(*//状态输出*)(*状态显示，容易造成指针容量不足*)
mov( ConveyorMotor.xEmpty AND NOT ConveyorMotor.xBusy , 0 , m_wStateWord);
mov( ConveyorMotor.xEmpty=0 , 							1 , m_wStateWord);
mov( ConveyorMotor.xBusy , 								2 , m_wStateWord);
mov( ConveyorMotor.xLimitAlarrm , 						3, 	m_wStateWord);
mov(ConveyorMotor.xOverWidthAlarm , 					4 , m_wStateWord);
mov( ConveyorMotor.xNotArriveAlarm , 					5 , m_wStateWord);
mov( ConveyorMotor.xUnloadAlarm, 						6 , m_wStateWord);
(*选择本线体后，将状态赋值给全局变量进行显示*)
mov( ConveyorMotor.diDeviceID=g_diDeviceIDSelect , m_wStateWord, g_iConveyorStatus );
END_FUNCTION_BLOCK

PROGRAM TCP
VAR
  m_ton1ReceiveHeartbeat : TON;
  m_t1RecHeartbeatCurrentTime : TIME;
  m_tonAutoClose : TON;
  m_xAutoClose : BOOL;
  m_tAutoCloseCurrentTime : TIME;
  m_tonReconnect : TON;
  m_xReconnect : BOOL;
  m_tReconnectCurrentTime : TIME;
  m_ton5ReceiveHeartbeat : TON;
  m_t5RecHeartbeatCurrentTime : TIME;
END_VAR
D220:=2;
m_tonReconnect(IN:= NOT SD1282.0 AND NOT SD1284.0 AND NOT m_xReconnect ,PT:=T#5s  ,Q:=m_xReconnect ,ET:=m_tReconnectCurrentTime);
SP_SOCOPEN(m_xReconnect  AND SD1288.A , "U0", K1 , D110 , M100);
SP_SOCSND( SM412 AND SD1282.0 , "U0" , K1 , D100, D220, M102 );
SP_SOCRCV( SD1282.0 AND SD1286.0 AND NOT M104 , "U0" , K1, D300 , D420 ,M104 );
m_tonAutoClose(IN:= SD1284.0 AND NOT SD1282.0 ,PT:=T#5s,Q:=m_xAutoClose ,ET:= m_tAutoCloseCurrentTime );
SP_SOCCLOSE( LDF(TRUE,SD1282.0) OR m_xAutoClose  , "U0" , K1, D120, M106 );
D221.F:=SM413;
m_ton1ReceiveHeartbeat(IN:=NOT LDP(TRUE, D421.F) ,PT:= t#5S ,Q:= g_xTcpFailed ,ET:= m_t1RecHeartbeatCurrentTime);
IF g_xTcpFailed THEN
	M104:=SM413;(*通讯失败有可能是接收模块没动作，重启接收模块*)
	D420:=0;
	D421:=0;
END_IF;

(*测试一下通信恢复功能*)
IF  g_xTcpFailed THEN
	SD1284.0:=SM414;
	SD414:=20;
END_IF;
END_PROGRAM

FUNCTION_BLOCK UConveyor
VAR
  iStep : INT;
END_VAR
VAR_IN_OUT
  ConveyorIOLeft : ConveyorIO;  (* U的左半边 *)
  ConveyorIORight : ConveyorIO;  (* U的右半边 *)
  ConveyorIODown : ConveyorIO;  (* U的下边一横 *)
  UConveyorIO : UConveyorIO;  (* 顶升,阻挡 *)
END_VAR
VAR
  m_xInitial : BOOL;
  m_tonCylinderOvertime : TON;  (* 气缸超时报警定时器 *)
  m_tCylinderOvertimeCurrent : TIME;
  m_tonExitBarDelay : TON;  (* 退出阻挡器延时 *)
  m_tExitBarDelay : TIME;
  m_xExitBarDelay : BOOL;
END_VAR
(*                                                                                                          
           

//*)
IF NOT m_xInitial THEN
	UConveyorIO.tSetOvertime:=T#5s;
	UConveyorIO.xExitEnable1:=1;
	UConveyorIO.xExitEnable2:=1;
	UConveyorIO.xExitEnable3:=1;
	m_xInitial:=1;
END_IF;
(*外部不用写ConveyorDown的开关，会自己根据来料的产品信息判断停哪个光电*)
IF UConveyorIO.iTask=1 AND ConveyorIODown.diDesConveyorIn=ConveyorIOLeft.diDeviceID THEN
	ConveyorIODown.xCWPresent:=ConveyorIOLeft.xCWPresent;
ELSIF UConveyorIO.iTask=1 AND ConveyorIODown.diDesConveyorIn=ConveyorIORight.diDeviceID THEN
	ConveyorIODown.xCWPresent:=ConveyorIORight.xCWPresent;
ELSE
	ConveyorIODown.xCWPresent:=ConveyorIOLeft.xCWPresent OR ConveyorIORight.xCWPresent;
END_IF;
(*这里判断什么时候直接放行，左右都不需要，也不是0，就放走*)
IF  NOT(ConveyorIODown.diDesConveyor=ConveyorIOLeft.diDeviceID 
		OR  ConveyorIODown.diDesConveyor=ConveyorIORight.diDeviceID 
		OR ConveyorIODown.diDesConveyor=0) THEN
	UConveyorIO.xPassEnable:=1;
ELSE
	UConveyorIO.xPassEnable:=0;
END_IF;	
IF g_xAuto THEN	
CASE UConveyorIO.iTask OF(*这个Task做抢占，可做LastTask保护*)
0:(*各种初始化，能自动去3*)
	ConveyorIODown.xLoad:=0;
	ConveyorIOleft.xLoad:=0;
	ConveyorIORight.xLoad:=0;
	ConveyorIODown.xUnload:=0;
	ConveyorIOLeft.xUnload:=0;
	ConveyorIORight.xUnload:=0;
	ConveyorIODown.xPutInto:=0;
	ConveyorIOLeft.xPutInto:=0;
	ConveyorIORight.xPutInto:=0;
	UConveyorIO.xExitBarCylinderRetract1:=0;
	UConveyorIO.xExitBarCylinderRetract2:=0;	
1:(*上料*)
	CASE iStep OF
	0:(*各种初始化，能自动去3*)
		ConveyorIODown.xLoad:=0;
		ConveyorIOleft.xLoad:=0;
		ConveyorIORight.xLoad:=0;
		ConveyorIODown.xUnload:=0;
		ConveyorIOLeft.xUnload:=0;
		ConveyorIORight.xUnload:=0;
		ConveyorIODown.xPutInto:=0;
		ConveyorIOLeft.xPutInto:=0;
		ConveyorIORight.xPutInto:=0;
		UConveyorIO.xExitBarCylinderRetract1:=0;
		UConveyorIO.xExitBarCylinderRetract2:=0;
		UConveyorIO.xBatteryError:=0;
		IF  NOT ConveyorIODown.xEmpty THEN
			iStep:=3;
		ELSE
			iStep:=1;
		END_IF;	
	1:(*顶升，等load*)
		IF UConveyorIO.xLiftCylinderExtendInit1 THEN
			UConveyorIO.xLiftCylinderExtend1:=1;
			UConveyorIO.xLiftCylinderRetract1:=0;
		ELSE
			UConveyorIO.xLiftCylinderExtend1:=0;
			UConveyorIO.xLiftCylinderRetract1:=1;
		END_IF;
		IF UConveyorIO.xLiftCylinderExtendInit2 THEN
			UConveyorIO.xLiftCylinderExtend2:=1;
			UConveyorIO.xLiftCylinderRetract2:=0;
			ELSE
			UConveyorIO.xLiftCylinderExtend2:=0;
			UConveyorIO.xLiftCylinderRetract2:=1;
		END_IF;
		IF 	((UConveyorIO.xLiftCylinderExtendInit1 AND UConveyorIO.xLiftCylinderExtendDetect1)
				OR (NOT UConveyorIO.xLiftCylinderExtendInit1 AND UConveyorIO.xLiftCylinderRetractDetect1))
			AND	((UConveyorIO.xLiftCylinderExtendInit2 AND UConveyorIO.xLiftCylinderExtendDetect2)
		   		OR (NOT UConveyorIO.xLiftCylinderExtendInit2 AND UConveyorIO.xLiftCylinderRetractDetect2))		
			AND	UConveyorIO.xEntryEnable1 THEN(*有上料请求1*)
		   	ConveyorIODown.xLoad:=1;
			iStep:=2;
		END_IF;
	2:(*Load完成*)(*去右臂时才需要阻挡放行,其他挡住*)
		UConveyorIO.xExitBarCylinderRetract1:=ConveyorIODown.diDesConveyorIn=ConveyorIORight.diDeviceID;
		IF NOT ConveyorIODown.xEmpty THEN
			ConveyorIODown.xLoad:=0;
			ConveyorIOLeft.xPutInto:=1;
			ConveyorIOright.xPutInto:=1;
			istep:=3;
		END_IF;
	3:(*顶升等Unload，这里等有了ExitEnable再顶升，因为可能有地方需要允许了再升降，比如倍速链*)
	IF (ConveyorIODown.diDesConveyor=ConveyorIOLeft.diDeviceID OR ConveyorIODown.diDesConveyor=ConveyorIORight.diDeviceID)
			AND	(UConveyorIO.xBatteryDetect1 OR UConveyorIO.xBatteryDetect2)(*在下面时检测*)
			AND UConveyorIO.xLiftCylinderRetractDetect1 AND UConveyorIO.xLiftCylinderRetractDetect2 THEN
			UConveyorIO.xBatteryError:=1;
		END_IF;	
		IF (ConveyorIODown.diDesConveyor=ConveyorIOLeft.diDeviceID AND UConveyorIO.xExitEnable2 AND NOT UConveyorIO.xBatteryError)THEN
			IF UConveyorIO.xLiftCylinderExtendInit1 THEN
				UConveyorIO.xLiftCylinderExtend1:=0;
				UConveyorIO.xLiftCylinderRetract1:=1;
			ELSE
				UConveyorIO.xLiftCylinderExtend1:=1;
				UConveyorIO.xLiftCylinderRetract1:=0;
			END_IF;
			IF(NOT UConveyorIO.xLiftCylinderExtendInit1 AND UConveyorIO.xLiftCylinderExtendDetect1)
				OR (UConveyorIO.xLiftCylinderExtendInit1 AND UConveyorIO.xLiftCylinderRetractDetect1)THEN
				iStep:=4;
			END_IF;
		END_IF;	
		IF (ConveyorIODown.diDesConveyor=ConveyorIORight.diDeviceID AND UConveyorIO.xExitEnable3 AND NOT UConveyorIO.xBatteryError)THEN
			IF UConveyorIO.xLiftCylinderExtendInit2 THEN
				UConveyorIO.xLiftCylinderExtend2:=0;
				UConveyorIO.xLiftCylinderRetract2:=1;
			ELSE
				UConveyorIO.xLiftCylinderExtend2:=1;
				UConveyorIO.xLiftCylinderRetract2:=0;
			END_IF;
			IF(NOT UConveyorIO.xLiftCylinderExtendInit2 AND UConveyorIO.xLiftCylinderExtendDetect2)
				OR (UConveyorIO.xLiftCylinderExtendInit2 AND UConveyorIO.xLiftCylinderRetractDetect2)THEN
				iStep:=4;
			END_IF;
		END_IF;	
		IF UConveyorIO.xPassEnable AND UConveyorIO.xExitEnable1 AND NOT UConveyorIO.xBatteryError THEN
			IF UConveyorIO.xLiftCylinderExtendInit1 THEN
				UConveyorIO.xLiftCylinderExtend1:=1;
				UConveyorIO.xLiftCylinderRetract1:=0;
			ELSE
				UConveyorIO.xLiftCylinderExtend1:=0;
				UConveyorIO.xLiftCylinderRetract1:=1;
			END_IF;
			IF UConveyorIO.xLiftCylinderExtendInit2 THEN
				UConveyorIO.xLiftCylinderExtend2:=0;
				UConveyorIO.xLiftCylinderRetract2:=1;
			ELSE
				UConveyorIO.xLiftCylinderExtend2:=1;
				UConveyorIO.xLiftCylinderRetract2:=0;
			END_IF;
			IF((UConveyorIO.xLiftCylinderExtendInit1 AND UConveyorIO.xLiftCylinderExtendDetect1)
					OR (NOT UConveyorIO.xLiftCylinderExtendInit1 AND UConveyorIO.xLiftCylinderRetractDetect1))
				AND((UConveyorIO.xLiftCylinderExtendInit2 AND UConveyorIO.xLiftCylinderExtendDetect2)
					OR (NOT UConveyorIO.xLiftCylinderExtendInit2 AND UConveyorIO.xLiftCylinderRetractDetect2))THEN
				UConveyorIO.xExitBarCylinderRetract1:=1;
				UConveyorIO.xExitBarCylinderRetract2:=1;
				iStep:=4;	
			END_IF;	
		END_IF;
	4:(*Unload完成，回0*)
			IF ConveyorIODown.diDesConveyor=ConveyorIOLeft.diDeviceID AND UConveyorIO.xExitEnable2 AND m_xExitBarDelay THEN
				ConveyorIOLeft.xUnloadCCW:=1;
				ConveyorIOLeft.xUnload:=1;
			ELSIF ConveyorIODown.diDesConveyor=ConveyorIORight.diDeviceID AND UConveyorIO.xExitEnable3 AND m_xExitBarDelay THEN
				ConveyorIORight.xUnloadCCW:=1;
				ConveyorIORight.xUnload:=1;
			ELSIF UConveyorIO.xPassEnable AND UConveyorIO.xExitEnable1 AND m_xExitBarDelay THEN
				ConveyorIODown.xUnload:=1;
			ELSE
				ConveyorIODown.xUnload:=0;
				ConveyorIOLeft.xUnload:=0;
				ConveyorIORight.xUnload:=0;
			END_IF;	
		IF ( (ConveyorIODown.diDesConveyor=ConveyorIOLeft.diDeviceID  AND LDF(TRUE,UConveyorIO.xExitEnable2))
		  OR(ConveyorIODown.diDesConveyor=ConveyorIORight.diDeviceID AND LDF(TRUE,UConveyorIO.xExitEnable3))
		  OR(UConveyorIO.xPassEnable AND LDF(TRUE,UConveyorIO.xExitEnable1)) )AND m_xExitBarDelay  THEN
			ConveyorIODown.xUnload:=0;
			ConveyorIOLeft.xUnload:=0;
			ConveyorIORight.xUnload:=0;
			ConveyorIODown.xPutInto:=1;
			ConveyorIOLeft.xPutInto:=1;
			ConveyorIORight.xPutInto:=1;
			UConveyorIO.xExitBarCylinderRetract1:=0;
			UConveyorIO.xExitBarCylinderRetract2:=0;
			iStep:=0;
		END_IF;
	END_CASE;
2:(*左下料*)
	CASE iStep OF
	0:(*各种初始化，能自动去3*)
		ConveyorIODown.xLoad:=0;
		ConveyorIOleft.xLoad:=0;
		ConveyorIORight.xLoad:=0;
		ConveyorIODown.xUnload:=0;
		ConveyorIOLeft.xUnload:=0;
		ConveyorIORight.xUnload:=0;
		ConveyorIODown.xPutInto:=0;
		ConveyorIOLeft.xPutInto:=0;
		ConveyorIORight.xPutInto:=0;
		UConveyorIO.xExitBarCylinderRetract1:=0;
		UConveyorIO.xExitBarCylinderRetract2:=0;
		UConveyorIO.xBatteryError:=0;
		IF  NOT ConveyorIODown.xEmpty THEN
			iStep:=3;
			ELSE
			iStep:=1;
		END_IF;	
	1:(*顶升，等load*)
		IF UConveyorIO.xLiftCylinderExtendInit1 THEN
			UConveyorIO.xLiftCylinderExtend1:=0;
			UConveyorIO.xLiftCylinderRetract1:=1;
			ELSE
			UConveyorIO.xLiftCylinderExtend1:=1;
			UConveyorIO.xLiftCylinderRetract1:=0;
		END_IF;
		IF ((NOT UConveyorIO.xLiftCylinderExtendInit1 AND UConveyorIO.xLiftCylinderExtendDetect1)
			OR ( UConveyorIO.xLiftCylinderExtendInit1 AND UConveyorIO.xLiftCylinderRetractDetect1))
			AND UConveyorIO.xEntryEnable2 THEN(*有上料请求1*)
		   	ConveyorIOLeft.xLoad:=1;
			iStep:=2;
		END_IF;
	2:(*Load完成*)
		IF NOT ConveyorIOLeft.xEmpty THEN
			ConveyorIOLeft.xLoad:=0;
			ConveyorIODown.xPutInto:=1;
			ConveyorIODown.diDesConveyor:=ConveyorIOLeft.diDesConveyor;
			istep:=3;
		END_IF;
	3:(*顶升等Unload，这里等有了ExitEnable再顶升，因为可能有地方需要允许了再升降，比如倍速链*)
		UConveyorIO.xExitBarCylinderRetract1:=1;
		UConveyorIO.xExitBarCylinderRetract2:=1;
		IF  UConveyorIO.xExitEnable1 THEN(*顶升共用一个汽缸得了*)
			IF UConveyorIO.xLiftCylinderExtendInit1 THEN
				UConveyorIO.xLiftCylinderExtend1:=1;
				UConveyorIO.xLiftCylinderRetract1:=0;
			ELSE
				UConveyorIO.xLiftCylinderExtend1:=0;
				UConveyorIO.xLiftCylinderRetract1:=1;
			END_IF;
		END_IF;
		IF UConveyorIO.xExitEnable1 THEN(*顶升共用一个汽缸得了*)
			IF(( UConveyorIO.xLiftCylinderExtendInit1 AND UConveyorIO.xLiftCylinderExtendDetect1)
				OR (NOT UConveyorIO.xLiftCylinderExtendInit1 AND UConveyorIO.xLiftCylinderRetractDetect1))THEN
				iStep:=4;
			END_IF;	
		END_IF;
	4:(*Unload完成，回0*)
		IF  UConveyorIO.xExitEnable1 AND m_xExitBarDelay THEN
			ConveyorIODown.xUnload:=1;
		ELSE
			ConveyorIODown.xUnload:=0;
		END_IF;	
		IF NOT UConveyorIO.xExitEnable1 AND m_xExitBarDelay   THEN
			ConveyorIODown.xUnload:=0;
			ConveyorIOLeft.xUnload:=0;
			ConveyorIORight.xUnload:=0;
			ConveyorIODown.xPutInto:=1;
			ConveyorIOLeft.xPutInto:=1;
			ConveyorIORight.xPutInto:=1;
			UConveyorIO.xExitBarCylinderRetract1:=0;
			UConveyorIO.xExitBarCylinderRetract2:=0;
			iStep:=0;
		END_IF;
	END_CASE;
3:(*上料到出口*)
	CASE iStep OF
	0:(*各种初始化，能自动去3*)
		ConveyorIODown.xLoad:=0;
		ConveyorIOleft.xLoad:=0;
		ConveyorIORight.xLoad:=0;
		ConveyorIODown.xUnload:=0;
		ConveyorIOLeft.xUnload:=0;
		ConveyorIORight.xUnload:=0;
		ConveyorIODown.xPutInto:=0;
		ConveyorIOLeft.xPutInto:=0;
		ConveyorIORight.xPutInto:=0;
		UConveyorIO.xExitBarCylinderRetract1:=0;
		UConveyorIO.xExitBarCylinderRetract2:=0;
		UConveyorIO.xBatteryError:=0;
		IF  NOT ConveyorIODown.xEmpty THEN
			iStep:=3;
		ELSE
			iStep:=1;
		END_IF;	
	1:(*顶升，等load*)
		IF UConveyorIO.xLiftCylinderExtendInit2 THEN
			UConveyorIO.xLiftCylinderExtend2:=0;
			UConveyorIO.xLiftCylinderRetract2:=1;
		ELSE
			UConveyorIO.xLiftCylinderExtend2:=1;
			UConveyorIO.xLiftCylinderRetract2:=0;
		END_IF;
		IF ((NOT UConveyorIO.xLiftCylinderExtendInit2 AND UConveyorIO.xLiftCylinderExtendDetect2)
			OR ( UConveyorIO.xLiftCylinderExtendInit2 AND UConveyorIO.xLiftCylinderRetractDetect2))
			AND UConveyorIO.xEntryEnable3 THEN(*有上料请求1*)
		   	ConveyorIORight.xLoad:=1;
			iStep:=2;
		END_IF;
	2:(*Load完成*)
		IF NOT ConveyorIORight.xEmpty THEN
			ConveyorIORight.xLoad:=0;
			ConveyorIODown.diDesConveyor:=ConveyorIORight.diDesConveyor;
			ConveyorIODown.xPutInto:=1;
			istep:=3;
		END_IF;
	3:(*顶升等Unload，这里等有了ExitEnable再顶升，因为可能有地方需要允许了再升降，比如倍速链*)
		UConveyorIO.xExitBarCylinderRetract2:=1;
		IF  UConveyorIO.xExitEnable1 THEN(*顶升共用一个汽缸得了*)
			IF UConveyorIO.xLiftCylinderExtendInit2 THEN
				UConveyorIO.xLiftCylinderExtend2:=1;
				UConveyorIO.xLiftCylinderRetract2:=0;
			ELSE
				UConveyorIO.xLiftCylinderExtend2:=0;
				UConveyorIO.xLiftCylinderRetract2:=1;
			END_IF;
		END_IF;
		IF UConveyorIO.xExitEnable1 THEN(*顶升共用一个汽缸得了*)
			IF(( UConveyorIO.xLiftCylinderExtendInit2 AND UConveyorIO.xLiftCylinderExtendDetect2)
				OR (NOT UConveyorIO.xLiftCylinderExtendInit2 AND UConveyorIO.xLiftCylinderRetractDetect2))THEN
				iStep:=4;
			END_IF;	
		END_IF;
	4:(*Unload完成，回0*)
		IF  UConveyorIO.xExitEnable1 AND m_xExitBarDelay THEN
			ConveyorIODown.xUnload:=1;
		ELSE
			ConveyorIODown.xUnload:=0;
		END_IF;	
		IF NOT UConveyorIO.xExitEnable1 AND m_xExitBarDelay  THEN
			ConveyorIODown.xUnload:=0;
			ConveyorIOLeft.xUnload:=0;
			ConveyorIORight.xUnload:=0;
			ConveyorIODown.xPutInto:=1;
			ConveyorIOLeft.xPutInto:=1;
			ConveyorIORight.xPutInto:=1;
			UConveyorIO.xExitBarCylinderRetract1:=0;
			UConveyorIO.xExitBarCylinderRetract2:=0;
			iStep:=0;
		END_IF;
	END_CASE;
END_CASE;(*iTask*)
m_tonExitBarDelay(IN:=iStep=4 ,PT:= T#1s ,Q:= m_xExitBarDelay ,ET:= m_tExitBarDelay);
END_IF;(*g_xAuto那个IF*)
(*复位程序*)
IF (g_xResetSingle AND  (g_diDeviceIDSelect=ConveyorIOLeft.diDeviceID 
						 OR g_diDeviceIDSelect=ConveyorIORight.diDeviceID
						 OR g_diDeviceIDSelect=ConveyorIODown.diDeviceID))
	OR LDP(TRUE,UConveyorIO.xLiftCylinderExtendInit1) 
	OR LDF(TRUE,UConveyorIO.xLiftCylinderExtendInit1) 
	OR LDP(TRUE,UConveyorIO.xPutInto)  THEN
	ConveyorIODown.xPutInto:=1;
	ConveyorIOLeft.xPutInto:=1;
	ConveyorIORight.xPutInto:=1;
	iStep:=0;
END_IF;
(*手动*)
IF g_xManual  THEN
	iStep:=0;
	ConveyorIODown.xLoad:=0;
	ConveyorIOleft.xLoad:=0;
	ConveyorIORight.xLoad:=0;
	ConveyorIODown.xUnload:=0;
	ConveyorIOLeft.xUnload:=0;
	ConveyorIORight.xUnload:=0;
	ConveyorIODown.xPutInto:=0;
	ConveyorIOLeft.xPutInto:=0;
	ConveyorIORight.xPutInto:=0;
	UConveyorIO.xBatteryError:=0;
	UConveyorIO.xLiftCylinderExtend1:=UConveyorIO.xLiftCylinderExtendButton1 AND NOT UConveyorIO.xLiftCylinderRetractButton1;
	UConveyorIO.xLiftCylinderRetract1:=UConveyorIO.xLiftCylinderRetractButton1 AND NOT UConveyorIO.xLiftCylinderExtendButton1;
	UConveyorIO.xLiftCylinderExtend2:=UConveyorIO.xLiftCylinderExtendButton2 AND NOT UConveyorIO.xLiftCylinderRetractButton2;
	UConveyorIO.xLiftCylinderRetract2:=UConveyorIO.xLiftCylinderRetractButton2 AND NOT UConveyorIO.xLiftCylinderExtendButton2;
	UConveyorIO.xExitBarCylinderRetract1:=UConveyorIO.xExitBarCylinderRetractButton1;
	UConveyorIO.xExitBarCylinderRetract2:=UConveyorIO.xExitBarCylinderRetractButton2;
END_IF;	
(*气缸超时报警*)
m_tonCylinderOvertime(IN:= (UConveyorIO.xLiftCylinderExtend1 AND NOT UConveyorIO.xLiftCylinderExtendDetect1) 
							OR  (UConveyorIO.xLiftCylinderRetract1 AND NOT UConveyorIO.xLiftCylinderRetractDetect1) 
							OR  (UConveyorIO.xLiftCylinderRetract2 AND NOT UConveyorIO.xLiftCylinderRetractDetect2) 
							OR  (UConveyorIO.xLiftCylinderRetract2 AND NOT UConveyorIO.xLiftCylinderRetractDetect2) ,
					PT:= UConveyorIO.tSetOvertime ,Q:=UConveyorIO.xOvertimeAlarm ,ET:=m_tCylinderOvertimeCurrent );
END_FUNCTION_BLOCK

FUNCTION ShuttleCarCurrentPosition
VAR_INPUT
  xPosition1 : BOOL;
  xPosition2 : BOOL;
  xPosition3 : BOOL;
END_VAR
(*//计算输送车当前位置的函数*)
IF xPosition1 THEN
	ShuttleCarCurrentPosition:=1;
END_IF;
IF xPosition2 THEN
	ShuttleCarCurrentPosition:=2;
END_IF;
IF xPosition3 THEN
	ShuttleCarCurrentPosition:=3;
END_IF;
END_FUNCTION

PROGRAM 批量复制专用
(*1线送出*)
	ConveyorIO401101.xUnload:=ConveyorIO40138.xEmpty AND LifterIO40203.iCurrentPos=2  AND X43 AND m_xPickDone[1];
	LifterIO40203.xMDIExe:=NOT ConveyorIO40138.xError AND NOT ConveyorIO401101.xError AND NOT ConveyorIO40131.xError;
	IF ConveyorIO40138.xEmpty THEN
		LifterIO40203.iDestinationPos:=2;
	ELSE
		LifterIO40203.iDestinationPos:=1;
	END_IF;		
	ConveyorIO40138.xLoad:=ConveyorIO401101.xNextRun;
	(*这里就不做抢占任务了，在下料条件里加上not busy信号得了。这样可能一个任务一直跑，所以可能有问题*)
	(*但是这样不用写任务，故障恢复容易些*)
	ConveyorIO40138.xUnload:=ConveyorIO40131.xEmpty AND LifterIO40203.iCurrentPos=1 AND X42
														AND NOT ConveyorIO40132.xBusy;(*未处于运行状态，表示没有在执行任务*)
	ConveyorIO40138.xUnloadCCW:=1;
	SwitchIO40312.xEntryEnable:=ConveyorIO40138.xNextRun;
	SwitchIO40312.xSwithEnable:=1;
	SwitchIO40312.xExitEnable:=ConveyorIO40133.xEmpty;
	(*ConveyorIO40134.xLoad:=ConveyorIO40132.xNextRun;
	ConveyorIO40134.xUnload:=ConveyorIO40133.xEmpty;*)
	ConveyorIO40133.xLoad:=ConveyorIO40132.xNextRun;
	ConveyorIO40133.xUnload:=D421.6;
	D221.6:=ConveyorIO40133.xNextRun;
	(*送出到出口大直线那里了*)
END_PROGRAM

FUNCTION_BLOCK Folder
VAR_IN_OUT
  FolderIO : FolderIO;
END_VAR
VAR
  m_xInitial : BOOL;
END_VAR
VAR_IN_OUT
  FolderConveyorIO : ConveyorIO;
END_VAR
VAR_GLOBAL RETAIN
  iFolderCount : INT;
END_VAR
VAR
  istep : INT;
  m_TONLoadDelay : TON;  (* 上料完成延时 *)
  m_xLoadDelay : BOOL;  (* 上料完成延时 *)
  m_tLoadDelay : TIME;  (* 上料完成延时 *)
  m_TONUpCylinderError : TON;
  m_tUpCylinderError : TIME;
  m_TONDownCylinderError : TON;
  m_tDownCylinderError : TIME;
  m_TONGrabCylinderError : TON;
  m_tGrabCylinderError : TIME;
END_VAR
VAR_INPUT
  i_xAuto : BOOL;  (* 自动 *)
  i_xManual : BOOL;  (* 手动 *)
END_VAR
(*叠盘机*)
(*李科远写的*)
(*初始化*)
IF NOT m_xInitial THEN
	FolderIO.i_iFloor:=3;
	FolderIO.i_tSetOvertime:=T#5S;
	
	m_xInitial:=1;
END_IF;
(*自动*)
FolderIO.o_xEntryPermit:=FolderConveyorIO.xEmpty;(*叠盘机的话，只要空了，就允许上料，拆盘则是拆完才允许*)
IF i_xAuto THEN
				m_TONLoadDelay(IN:= NOT FolderConveyorIO.xEmpty,
													PT:= T#100MS,
													Q:=m_xLoadDelay,
													ET:=m_tLoadDelay);
	CASE istep OF
		0:(*各种初始化*)
			FolderConveyorIO.xLoad:=0;
			FolderConveyorIO.xUnload:=0;
			FolderConveyorIO.xPutInto:=0;
			IF 0 AND  FolderConveyorIO.xEmpty THEN
				istep:=1;(*空着就去1上料*)
			END_IF;	
			IF 0 AND    m_xLoadDelay  THEN(*if 有料*)
				IF  FolderIO.i_xCylinderDownExtendDetect  AND FolderIO.i_xCylinderUpExtendDetect  THEN(*if 在下层*)
					IF iFolderCount=FolderIO.i_iFloor THEN(*if 是最后一次*)
						istep:=7;
					ELSE(*不是最后一次去5，是就去7*)
						istep:=5;
					END_IF;(*if 是最后一次*)	
				ELSE(*不在下层去2*)
				istep:=2;
				END_IF;	(*if 在下层*)			
			END_IF;(*if 有料*)
			
		1:(*上料*)
			IF FolderIO.i_xEntryEnable THEN
				FolderConveyorIO.xLoad:=1;
			ELSE
				FolderConveyorIO.xLoad:=0;
			END_IF;(*not Empty了等个延时*)	

			IF 0 AND   m_xLoadDelay  AND (iFolderCount>0 AND iFolderCount<FolderIO.i_iFloor) THEN
				istep:=2;
			ELSIF 0 AND   m_xLoadDelay AND iFolderCount=0 THEN(*=0表示是第一次，第一次直接抓紧上升*)
				istep:=5;	
			END_IF;	
		2:(*下降，到2层位置*)
				FolderIO.o_xCylinderUpRetract:=0;
				FolderIO.o_xCylinderUpExtend:=1;
				FolderIO.o_xCylinderDownRetract:=1;
				FolderIO.o_xCylinderDownExtend:=0;
				IF 0 AND   FolderIO.i_xCylinderUpExtendDetect AND NOT FolderIO.i_xCylinderDownExtendDetect THEN
					istep:=3;
				END_IF;
		3:	(*松开夹爪*)
			IF FolderConveyorIO.xCWPresent AND NOT FolderConveyorIO.xEmpty THEN(*有感应到才松开*)
				FolderIO.o_xCylinderGrabExtend:=0;
				FolderIO.o_xCylinderGrabRetract:=1;
				IF 0 AND   FolderIO.i_xCylinderGrabRetractDetect THEN
					IF iFolderCount=FolderIO.i_iFloor-1 THEN
						iFolderCount:=FolderIO.i_iFloor;(*最后一次到这里就刷新计数，方便故障恢复*)
					END_IF;	
					istep:=4;
				END_IF;	
			END_IF;	
		4:(*再下降，去1层*)
				FolderIO.o_xCylinderUpRetract:=0;
				FolderIO.o_xCylinderUpExtend:=1;
				FolderIO.o_xCylinderDownRetract:=0;
				FolderIO.o_xCylinderDownExtend:=1;
				IF 0 AND   FolderIO.i_xCylinderDownExtendDetect  AND FolderIO.i_xCylinderUpExtendDetect  THEN
					IF iFolderCount<FolderIO.i_iFloor-1 THEN
						istep:=5;
					ELSE
						istep:=7;
					END_IF;	
				END_IF;		
		5:(*抓紧*)
			IF FolderIO.i_xCylinderDownExtendDetect  AND FolderIO.i_xCylinderUpExtendDetect  THEN
				FolderIO.o_xCylinderGrabExtend:=1;
				FolderIO.o_xCylinderGrabRetract:=0;
				IF 0 AND   FolderIO.i_xCylinderGrabExtendDetect THEN
					iFolderCount:=iFolderCount+1;
					istep:=6;
				END_IF;	
			END_IF;		
		6:(*上升到3层*)
			FolderIO.o_xCylinderUpRetract:=1;
			FolderIO.o_xCylinderUpExtend:=0;
			FolderIO.o_xCylinderDownRetract:=1;
			FolderIO.o_xCylinderDownExtend:=0;
			IF 0 AND   FolderIO.i_xCylinderDownRetractDetect AND FolderIO.i_xCylinderUpRetractDetect THEN
				FolderConveyorIO.xPutInto:=1;(*刷新成Empty的*)
				istep:=0;
			END_IF;
		7:(*下料*)	
				IF	FolderIO.i_xExitEnable AND FolderIO.i_xCylinderGrabRetractDetect	THEN(*保证不会挂到叉手*)
				FolderConveyorIO.xUnload:=1;
			ELSE
				FolderConveyorIO.xPutInto:=1;(*刷新成Empty的*)
				FolderConveyorIO.xUnload:=0;
			END_IF;	
			IF 0 AND   FolderConveyorIO.xEmpty THEN(*确保空了才回0，不然还在这里等Unload信号*)
				iFolderCount:=0;
				istep:=0;
			END_IF;	 
		END_CASE;
END_IF;(*g_xAuto那个*)	
(*手动控制气缸动作*)
		IF i_xManual THEN
			FolderIO.o_xCylinderGrabExtend:=	FolderIO.i_xCylinderGrabExtendButton;	
			FolderIO.o_xCylinderGrabRetract:=	FolderIO.i_xCylinderGrabRetractButton;	
			FolderIO.o_xCylinderUpExtend:=		FolderIO.i_xCylinderUpExtendButton;	
			FolderIO.o_xCylinderUpRetract:=		FolderIO.i_xCylinderUpRetractButton;	
			FolderIO.o_xCylinderDownExtend:=	FolderIO.i_xCylinderDownExtendButton;	
			FolderIO.o_xCylinderDownRetract:=	FolderIO.i_xCylinderDownRetractButton;		
		END_IF;
		
		(*气缸超时未到达报警，可能是没气儿漏气，也可能是开关坏了，或者气缸被卡住了*)
		m_TONGrabCylinderError(IN:= (FolderIO.o_xCylinderGrabExtend AND NOT FolderIO.i_xCylinderGrabExtendDetect) 
																OR  (FolderIO.o_xCylinderGrabRetract AND NOT FolderIO.i_xCylinderGrabRetractDetect) ,
															PT:= FolderIO.i_tSetOvertime ,Q:= FolderIO.o_xGrabCylinderError,ET:= m_tGrabCylinderError);
		m_TONDownCylinderError(IN:= (FolderIO.o_xCylinderDownExtend AND NOT FolderIO.i_xCylinderDownExtendDetect) 
																OR  (FolderIO.o_xCylinderDownRetract AND NOT FolderIO.i_xCylinderDownRetractDetect) ,
															PT:= FolderIO.i_tSetOvertime ,Q:= FolderIO.o_xDownCylinderError,ET:= m_tDownCylinderError);
		m_TONUpCylinderError(IN:= (FolderIO.o_xCylinderUpExtend AND NOT FolderIO.i_xCylinderUpExtendDetect) 
																OR  (FolderIO.o_xCylinderUpRetract AND NOT FolderIO.i_xCylinderUpRetractDetect) ,
															PT:= FolderIO.i_tSetOvertime ,Q:= FolderIO.o_xUpCylinderError,ET:= m_tUpCylinderError);
END_FUNCTION_BLOCK

FUNCTION_BLOCK DivideFolder
VAR_IN_OUT
  FolderIO : FolderIO;
  FolderConveyorIO : ConveyorIO;
END_VAR
VAR_GLOBAL RETAIN
  iFolderCount : INT;
END_VAR
VAR
  m_xInitial : BOOL;
  istep : INT;
  m_TONLoadDelay : TON;  (* 上料完成延时 *)
  m_xLoadDelay : BOOL;  (* 上料完成延时 *)
  m_tLoadDelay : TIME;  (* 上料完成延时 *)
  m_TONUpCylinderError : TON;
  m_tUpCylinderError : TIME;
  m_TONDownCylinderError : TON;
  m_tDownCylinderError : TIME;
  m_TONGrabCylinderError : TON;
  m_tGrabCylinderError : TIME;
END_VAR
(*叠盘机*)
(*初始化*)
IF NOT m_xInitial THEN
	FolderIO.i_iFloor:=3;
	FolderIO.i_tSetOvertime:=T#5S;
	
	m_xInitial:=1;
END_IF;
(*自动*)
IF g_xAuto THEN
	FolderIO.o_xEntryPermit:=iFolderCount=0 AND FolderConveyorIO.xEmpty;(*空了且数量为0了，才准上料*)
	m_TONLoadDelay(IN:= NOT FolderConveyorIO.xEmpty,
											PT:= T#100MS,
											Q:=m_xLoadDelay,
											ET:=m_tLoadDelay);
	CASE istep OF
		0:(*各种初始化*)
			FolderConveyorIO.xLoad:=0;
			FolderConveyorIO.xUnload:=0;
			FolderConveyorIO.xPutInto:=0;
			IF FolderConveyorIO.xEmpty THEN(*空的情况，0时上料，其他走流程*)
				IF iFolderCount=0  THEN
					istep:=1; 					
				ELSE 
					istep:=2;
				END_IF;	
			END_IF;		
			IF m_xLoadDelay THEN
				 IF FolderIO.i_xCylinderDownExtendDetect  AND FolderIO.i_xCylinderUpExtendDetect  THEN
					istep:=3;(*如果在下层执行3*)
				ELSIF FolderIO.i_xCylinderDownRetractDetect AND FolderIO.i_xCylinderUpRetractDetect THEN
					istep:=7;(*如果在上层执行下料过程*)
				 ELSE 
				 	istep:=5;(*如果在中层执行夹紧缩回流程*)
				END_IF;		
			END_IF;
		1:(*上料*)
			IF FolderIO.i_xEntryEnable THEN
				FolderConveyorIO.xLoad:=1;
			ELSE
				FolderConveyorIO.xLoad:=0;
			END_IF;(*not Empty了等个延时*)	

			IF m_xLoadDelay THEN
				iFolderCount:=FolderIO.i_iFloor;
				istep:=5;(**上料肯定是第一次才上料，所以必然去5，抓紧上升*)
			END_IF;	
		2:(*下降，到1层位置*)
				FolderIO.o_xCylinderUpRetract:=0;
				FolderIO.o_xCylinderUpExtend:=1;
				FolderIO.o_xCylinderDownRetract:=0;
				FolderIO.o_xCylinderDownExtend:=1;
				IF FolderIO.i_xCylinderDownExtendDetect AND FolderIO.i_xCylinderUpExtendDetect THEN
					istep:=3;
				END_IF;
		3:	(*松开夹爪*)
			IF FolderIO.i_xCylinderDownExtendDetect AND FolderIO.i_xCylinderUpExtendDetect THEN
				FolderIO.o_xCylinderGrabExtend:=0;
				FolderIO.o_xCylinderGrabRetract:=1;
			END_IF;
			IF FolderIO.i_xCylinderGrabRetractDetect THEN
				IF iFolderCount=1 THEN(*最后一次到这里就刷新数据，方便复位*)
					iFolderCount:=0;
				END_IF;	
				istep:=4;
			END_IF;	
		4:(*再上升到2层*)
				FolderIO.o_xCylinderUpRetract:=0;
				FolderIO.o_xCylinderUpExtend:=1;
				FolderIO.o_xCylinderDownRetract:=1;
				FolderIO.o_xCylinderDownExtend:=0;
				IF FolderIO.i_xCylinderDownRetractDetect  AND FolderIO.i_xCylinderUpExtendDetect  THEN
					IF iFolderCount=1 THEN(*最后一次到此为止，升到2层就算完成*)
						istep:=7;
					ELSE	(*其他都走正常流程*)
						istep:=5;
					END_IF;		
				END_IF;		
		5:(*抓紧*)
			IF FolderIO.i_xCylinderDownRetractDetect  AND FolderIO.i_xCylinderUpExtendDetect  THEN
				FolderIO.o_xCylinderGrabExtend:=1;
				FolderIO.o_xCylinderGrabRetract:=0;
				IF FolderIO.i_xCylinderGrabExtendDetect THEN
					istep:=6;
				END_IF;	
			END_IF;		
		6:(*上升到3层*)
			FolderIO.o_xCylinderUpRetract:=1;
			FolderIO.o_xCylinderUpExtend:=0;
			FolderIO.o_xCylinderDownRetract:=1;
			FolderIO.o_xCylinderDownExtend:=0;
			IF FolderIO.i_xCylinderDownRetractDetect AND FolderIO.i_xCylinderUpRetractDetect THEN
				FolderConveyorIO.xPutInto:=1;
				istep:=7;
			END_IF;
		7:(*下料*)	
			IF	FolderIO.i_xExitEnable	
				AND FolderIO.i_xCylinderDownExtendDetect (*通过这些保证我没有挂到叉手*)
				AND FolderIO.i_xCylinderUpExtendDetect  
				AND FolderIO.i_xCylinderGrabRetractDetect	THEN
				FolderConveyorIO.xUnload:=1;
			ELSE
				FolderConveyorIO.xPutInto:=1;
				FolderConveyorIO.xUnload:=0;
			END_IF;	
			IF FolderConveyorIO.xEmpty THEN
			FolderConveyorIO.xPutInto:=0;
				IF iFolderCount>1 THEN
					iFolderCount:=iFolderCount-1;					
					istep:=2;
				ELSE
					istep:=0;
				END_IF;	
			END_IF;		
		END_CASE;
END_IF;(*g_xAuto那个*)	
(*手动控制气缸动作*)
		IF g_xManual THEN
			FolderIO.o_xCylinderGrabExtend:=	FolderIO.i_xCylinderGrabExtendButton;	
			FolderIO.o_xCylinderGrabRetract:=	FolderIO.i_xCylinderGrabRetractButton;	
			FolderIO.o_xCylinderUpExtend:=		FolderIO.i_xCylinderUpExtendButton;	
			FolderIO.o_xCylinderUpRetract:=		FolderIO.i_xCylinderUpRetractButton;	
			FolderIO.o_xCylinderDownExtend:=	FolderIO.i_xCylinderDownExtendButton;	
			FolderIO.o_xCylinderDownRetract:=	FolderIO.i_xCylinderDownRetractButton;		
		END_IF;
		
		(*气缸超时未到达报警，可能是没气儿漏气，也可能是开关坏了，或者气缸被卡住了*)
		m_TONGrabCylinderError(IN:= (FolderIO.o_xCylinderGrabExtend AND NOT FolderIO.i_xCylinderGrabExtendDetect) 
																OR  (FolderIO.o_xCylinderGrabRetract AND NOT FolderIO.i_xCylinderGrabRetractDetect) ,
															PT:= FolderIO.i_tSetOvertime ,Q:= FolderIO.o_xGrabCylinderError,ET:= m_tGrabCylinderError);
		m_TONDownCylinderError(IN:= (FolderIO.o_xCylinderDownExtend AND NOT FolderIO.i_xCylinderDownExtendDetect) 
																OR  (FolderIO.o_xCylinderDownRetract AND NOT FolderIO.i_xCylinderDownRetractDetect) ,
															PT:= FolderIO.i_tSetOvertime ,Q:= FolderIO.o_xDownCylinderError,ET:= m_tDownCylinderError);
		m_TONUpCylinderError(IN:= (FolderIO.o_xCylinderUpExtend AND NOT FolderIO.i_xCylinderUpExtendDetect) 
																OR  (FolderIO.o_xCylinderUpRetract AND NOT FolderIO.i_xCylinderUpRetractDetect) ,
															PT:= FolderIO.i_tSetOvertime ,Q:= FolderIO.o_xUpCylinderError,ET:= m_tUpCylinderError);
END_FUNCTION_BLOCK

FUNCTION_BLOCK ConveyorCommunication
VAR_IN_OUT
  ConveyorIO : ConveyorIO;
  CommunicationIO : CommunicationIO;
END_VAR
VAR_OUTPUT
  o_iErrorNub : INT;  (* 错误代码 *)
END_VAR
VAR
  o_xReqSuccess : BOOL;  (* 请求成功 *)
  m_xInitial : BOOL;  (* 初始化 *)
  o_xError : BOOL;  (* 通信数据错误 *)
END_VAR
(********************************************************************************)
(*
DB1区(PC->PLC)15个字		
"字(16位）序号
(从1开始)"			功能描述											具体参数解释
1					请求确认	"										1：复位
				 														2：读码(入库申请）成功
				 														3：取放货完成 
																		4：旋转
																		5：不旋转
																		101：条码空
																		102：条码规则校验失败
																		103：步号校验失败
																		104：无库位可用 
"
2	预留	
3	预留	
4	预留	
5	预留	
6	读写标志位	"														1：写入数据
																		2：读数据完成"
7	任务处理标志	"														１：复位
																		２：完成"
8	命令字	"
																		21-送出（任务起点与终点不同，即向下一台输送机移载）
																		22：叠盘
"
9	任务号	"															1~65535唯一任务标识"
10	目标设备号															只有送出任务才有效
11		
12	筐码后4位	
				

DB2区(PLC->PC)15个字			
"字(16位）序号
(从1开始)"	功能描述	具体参数解释	
1	请求状态	"１：复位
２：请求"	实时状态，没有时序交互
2	强制入库(预留）	"１：复位
２：强制入库"	
3	预留(叠盘数量）	只对叠盘工位有效	
4	预留		
5			
6	读写标志位	"1：写入数据
2：读数据完成"	"有交互
时序"
7	设备状态	"1:空闲
2：工作中
3:任务完成（只有目标设备才会报任务完成）
４：故障"	
8	任务号	1~65535唯一任务标识，当输送任务执行完成后，将PC下发的任务号上报	
9	筐码后4位		
10	预留		
11			
			





2018.8.3 YAO 1.0
*)
(********************************************************************************)
(*如果外部不设置，就认为没有额外条件，有料就请求*)
IF NOT m_xInitial THEN
		CommunicationIO.i_xExtraCondition:=1;
		CommunicationIO.i_xExportConveyor:=0;
		m_xInitial:=1;
END_IF;
(*//有料状态*)
IF ConveyorIO.xEmpty THEN
	CommunicationIO.o_iEmptyPLCPC:=1;
	CommunicationIO.o_iRequestPLCPC:=1;(*无料撤销请求*)
	ELSE
	CommunicationIO.o_iEmptyPLCPC:=2;
END_IF;

(*//请求状态*)
(*入库段线体*)
IF CommunicationIO.i_xExportConveyor=0 THEN
(*非终点设备，满足条件才发请求，否则不发*)
		IF NOT ConveyorIO.xEmpty AND CommunicationIO.i_xExtraCondition THEN
			CommunicationIO.o_iRequestPLCPC:=2;
		ELSE
			CommunicationIO.o_iRequestPLCPC:=1;
		END_IF;
ELSIF CommunicationIO.i_xImportConveyor THEN
	IF ConveyorIO.diDesConveyor = ConveyorIO.diDeviceID THEN(*非终点设备，满足条件才发请求，否则不发*)
		IF NOT ConveyorIO.xEmpty AND CommunicationIO.i_xExtraCondition THEN
			CommunicationIO.o_iRequestPLCPC:=2;
		ELSE
			CommunicationIO.o_iRequestPLCPC:=1;
		END_IF;
	END_IF;
ELSE
		IF ConveyorIO.xEmpty AND CommunicationIO.i_xExtraCondition THEN
			CommunicationIO.o_iRequestPLCPC:=2;
		ELSE
			CommunicationIO.o_iRequestPLCPC:=1;
		END_IF;
END_IF;	
(*出库段线体*)
(*//请求确认*)
CASE CommunicationIO.i_iResponsPCPLC OF 
	0:;
	1:;(*//复位*)
	2:(*//读码（入库申请）成功*)
	o_xReqSuccess:=1;
	3:(*//取放货完成*)
	ConveyorIO.xPutInto:=1; 
	4:(*//旋转*)
	o_xReqSuccess:=1;
	ConveyorIO.xPutInto:=1; 
	5:(*//不旋转*)
	o_xReqSuccess:=1;
	ConveyorIO.xPutInto:=1; 
	101:(*//条码空*)
	o_iErrorNub:=101;
	o_xError:=1;
	102:(*//条码规则检验失败*)
	o_iErrorNub:=102;
	o_xError:=1;
	103:(*//步号校验失败*)
	o_iErrorNub:=103;
	o_xError:=1;
	104:(*//无库位可用*)
	o_iErrorNub:=104;
	o_xError:=1;
	105:(*//路径选择失败*)
	o_iErrorNub:=105;
	o_xError:=1;
	106:(*//控制ID错误*)
	o_iErrorNub:=106;
	o_xError:=1;
	107:(*//叠盘计数不一致*)
	o_iErrorNub:=107;
	o_xError:=1;
END_CASE;
(*IF LDP(TRUE,CommunicationIO.i_iResponsPCPLC=3
			OR CommunicationIO.i_iResponsPCPLC =4
			OR CommunicationIO.i_iResponsPCPLC =5 ) THEN
	ConveyorIO.xPutInto:=1;
END_IF;*)
IF LDP(TRUE,CommunicationIO.i_iResponsPCPLC <> 3
			AND CommunicationIO.i_iResponsPCPLC <>4
			AND CommunicationIO.i_iResponsPCPLC <>5 ) THEN
	ConveyorIO.xPutInto:=0;
END_IF;
IF CommunicationIO.i_iResponsPCPLC <> 2 
	AND CommunicationIO.i_iResponsPCPLC <>4
	AND CommunicationIO.i_iResponsPCPLC <>5 THEN
	o_xReqSuccess:=0;
END_IF;
IF CommunicationIO.i_iResponsPCPLC < 100 THEN
	o_iErrorNub:=0;
	o_xError:=0;
END_IF;

(*//读写标志位写入数据*)
IF ConveyorIO.diDesConveyor<>ConveyorIO.diDeviceID THEN
	IF LDP(TRUE,CommunicationIO.i_iReadWriteFlagPCPLC = 1) THEN
		ConveyorIO.iTaskID := CommunicationIO.i_iTaskIDPCPLC;
		ConveyorIO.diDesConveyor := CommunicationIO.i_diDestinationDevicePCPLC;
		ConveyorIO.iProductCategory :=CommunicationIO.i_iProductIDPCPLC;
	END_IF;
END_IF;
(*//数据校验，并返回握手信号*)
IF CommunicationIO.i_iReadWriteFlagPCPLC = 1 
	AND ConveyorIO.iTaskID<>0
	AND ConveyorIO.diDesConveyor<>0 
	(*AND ConveyorIO.iProductCategory<>0 *)
	THEN
	CommunicationIO.o_iReadWriteFlagPLCPC:=2;
	(*处理标志位为2时，返回一个2*)
	ELSIF CommunicationIO.i_iTaskProcessFlagPCPLC=2 THEN
		CommunicationIO.o_iReadWriteFlagPLCPC:=2;
	ELSE
	CommunicationIO.o_iReadWriteFlagPLCPC:=1;
END_IF;

(*//数据校验*)
IF CommunicationIO.i_iReadWriteFlagPCPLC = 1 
	AND (ConveyorIO.iTaskID<>0
	OR ConveyorIO.diDesConveyor<>0 )
	(*OR ConveyorIO.iProductCategory<>0) *)
	THEN
	o_iErrorNub:=50;(*//任务数据不完整*)
END_IF;
(*//设备状态*)
IF ConveyorIO.diDesConveyor = ConveyorIO.diDeviceID 
		AND (ldp(TRUE,NOT ConveyorIO.xEmpty AND CommunicationIO.i_xExtraCondition)
		OR (g_diDeviceIDSelect=ConveyorIO.diDeviceID AND ldp(TRUE,g_xInsertTask)))(*插入任务时，同时报一次完成*)
		THEN(*//目标地址=当前地址，表示是终点设备，有料就上传数据，报完成*)
	CommunicationIO.o_iDeviceStatusPLCPC:=3;(*//任务完成*)
	CommunicationIO.o_iProductIDPLCPC:=ConveyorIO.iProductCategory;(*//条码后四位上传*)
	CommunicationIO.o_iTaskIDPLCPC:=ConveyorIO.iTaskID;(*//任务号上传*)
	CommunicationIO.o_iRequestPLCPC:=2;(*发送入库请求*)
ELSIF ConveyorIO.diDesConveyor = ConveyorIO.diDeviceID AND LDp(TRUE,CommunicationIO.i_iTaskProcessFlagPCPLC=1)	
	THEN	(*//目标地址=当前地址，表示是终点设备，上位机给完成信号，就复位信号*)
	CommunicationIO.o_iDeviceStatusPLCPC:=1;
	CommunicationIO.o_iProductIDPLCPC:=0;(*//条码号复位*)
	CommunicationIO.o_iTaskIDPLCPC:=0;(*//任务号复位*)
ELSIF 	ConveyorIO.diDesConveyor <>ConveyorIO.diDeviceID AND (ConveyorIO.xEmpty OR (NOT ConveyorIO.xEmpty AND   CommunicationIO.i_xExtraCondition)) THEN(*非终点设备，无料就复位*)
	CommunicationIO.o_iDeviceStatusPLCPC:=1;
ELSIF ConveyorIO.xBusy THEN
	CommunicationIO.o_iDeviceStatusPLCPC:=2;(*//工作中*)
ELSIF ConveyorIO.xError THEN
	CommunicationIO.o_iDeviceStatusPLCPC:=4;(*//故障*)	
END_IF;
IF NOT g_xAuto THEN
	CommunicationIO.o_iDeviceStatusPLCPC:=0;
	CommunicationIO.o_iEmptyPLCPC:=0;
	CommunicationIO.o_iFolderNumberPLCPC:=0;
	CommunicationIO.o_iForceInportPLCPC:=0;
	CommunicationIO.o_iProductIDPLCPC:=0;
	CommunicationIO.o_iReadWriteFlagPLCPC:=0;
	CommunicationIO.o_iRequestPLCPC:=0;
	CommunicationIO.o_iTaskIDPLCPC:=0;
END_IF;
END_FUNCTION_BLOCK

PROGRAM START
IF g_xReset THEN
	SM50:=1;
	ELSE
	SM50:=0;
END_IF;
CASE g_iState OF
	0: (*手动*)
	g_xManual:=1;
	g_xAuto:=0;	
	g_xStackLampAmber:=1;
	g_xStackLampGreen:=0;
	g_xRemoteAuto:=0;
	g_xAutoLamp:=0;
	1:(*自动*)
	g_xManual:=0;
	g_xAuto:=1;
	g_xStackLampGreen:=1;
	g_xStackLampAmber:=0;
	g_xRemoteAuto:=0;
	g_xAutoLamp:=1;
	2:	(*远程自动*)
	g_xRemoteAuto:=1;
	g_xStackLampGreen:=1;
	g_xStackLampAmber:=0;
	g_xAuto:=0;
	g_xManual:=0;
	g_xAutoLamp:=0;
	3:(*自动未启动*)
	g_xRemoteAuto:=1;
	g_xStackLampGreen:=SM412;
	g_xStackLampAmber:=0;
	g_xAuto:=0;
	g_xManual:=0;	
	g_xAutoLamp:=0;
END_CASE;

IF g_xAutoSwitch AND g_xAutoStart  THEN  
	g_iState:=1;
END_IF;

IF g_xAutoSwitch AND (g_iState<>1 OR NOT g_xStop)  THEN  
	g_iState:=3;
END_IF;

g_xStackLampRed:=g_xAlarm AND SM412;
g_xBuzzer:=g_xAlarm AND SM412 AND NOT g_xMute;

IF LDF(TRUE,g_xAlarm) THEN
	g_xMute:=0;
END_IF;

IF NOT g_xAutoSwitch  OR g_xEStop=0 THEN 
	g_iState:=0;
END_IF;
IF g_xRemoteAutoStart THEN
	g_iState:=2;
END_IF;
IF g_xPause AND SM412 THEN
	g_xStackLampGreen:=0;
	g_xStackLampAmber:=0;
END_IF;
END_PROGRAM
